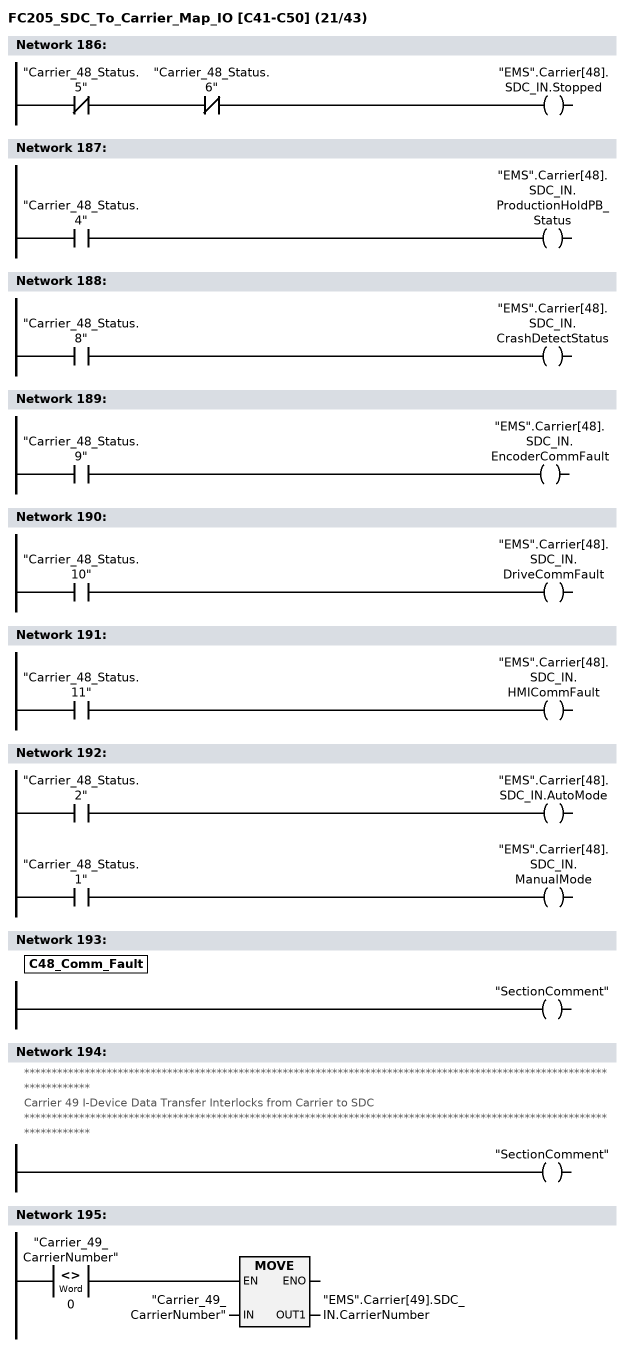
   RUNG wire#powerrail
      I_Contact( "Carrier_48_Status.5" )
      I_Contact( "Carrier_48_Status.6" )
      Coil( "EMS".Carrier[48].SDC_IN.Stopped )
   END_RUNG
   // the same network as SCL:
   "EMS".Carrier[48].SDC_IN.Stopped := NOT "Carrier_48_Status.5" AND NOT "Carrier_48_Status.6";
END_REGION

REGION Network 187
   RUNG wire#powerrail
      Contact( "Carrier_48_Status.4" )
      Coil( "EMS".Carrier[48].SDC_IN.ProductionHoldPB_Status )
   END_RUNG
   // the same network as SCL:
   "EMS".Carrier[48].SDC_IN.ProductionHoldPB_Status := "Carrier_48_Status.4";
END_REGION

REGION Network 188
   RUNG wire#powerrail
      Contact( "Carrier_48_Status.8" )
      Coil( "EMS".Carrier[48].SDC_IN.CrashDetectStatus )
   END_RUNG
   // the same network as SCL:
   "EMS".Carrier[48].SDC_IN.CrashDetectStatus := "Carrier_48_Status.8";
END_REGION

REGION Network 189
   RUNG wire#powerrail
      Contact( "Carrier_48_Status.9" )
      Coil( "EMS".Carrier[48].SDC_IN.EncoderCommFault )
   END_RUNG
   // the same network as SCL:
   "EMS".Carrier[48].SDC_IN.EncoderCommFault := "Carrier_48_Status.9";
END_REGION

REGION Network 190
   RUNG wire#powerrail
      Contact( "Carrier_48_Status.10" )
      Coil( "EMS".Carrier[48].SDC_IN.DriveCommFault )
   END_RUNG
   // the same network as SCL:
   "EMS".Carrier[48].SDC_IN.DriveCommFault := "Carrier_48_Status.10";
END_REGION

REGION Network 191
   RUNG wire#powerrail
      Contact( "Carrier_48_Status.11" )
      Coil( "EMS".Carrier[48].SDC_IN.HMICommFault )
   END_RUNG
   // the same network as SCL:
   "EMS".Carrier[48].SDC_IN.HMICommFault := "Carrier_48_Status.11";
END_REGION

REGION Network 192
   RUNG wire#powerrail
      Contact( "Carrier_48_Status.2" )
      Coil( "EMS".Carrier[48].SDC_IN.AutoMode )
   END_RUNG
   RUNG wire#powerrail
      Contact( "Carrier_48_Status.1" )
      Coil( "EMS".Carrier[48].SDC_IN.ManualMode )
   END_RUNG
   // the same network as SCL:
   "EMS".Carrier[48].SDC_IN.AutoMode := "Carrier_48_Status.2";
   "EMS".Carrier[48].SDC_IN.ManualMode := "Carrier_48_Status.1";
END_REGION

REGION Network 193
   Label( C48_Comm_Fault )
   RUNG wire#powerrail
      Coil( "SectionComment" )
   END_RUNG
   // the same network as SCL:
   C48_Comm_Fault:
   "SectionComment" := TRUE;
END_REGION

REGION Network 194
   // **********************************************************************************************************************
   // 
   // Carrier 49 I-Device Data Transfer Interlocks from Carrier to SDC
   // 
   // **********************************************************************************************************************
   RUNG wire#powerrail
      Coil( "SectionComment" )
   END_RUNG
   // the same network as SCL:
   "SectionComment" := TRUE;
END_REGION

REGION Network 195
   RUNG wire#powerrail
      { S7_Templates := "SrcType := Word" } NE_Contact(in1 := "Carrier_49_CarrierNumber", in2 := 0)
      Move(in := "Carrier_49_CarrierNumber", out1 => "EMS".Carrier[49].SDC_IN.CarrierNumber)
   END_RUNG
   // the same network as SCL:
   IF "Carrier_49_CarrierNumber" <> 0 THEN
       "EMS".Carrier[49].SDC_IN.CarrierNumber := "Carrier_49_CarrierNumber";
   END_IF;
END_REGION

REGION Network 196
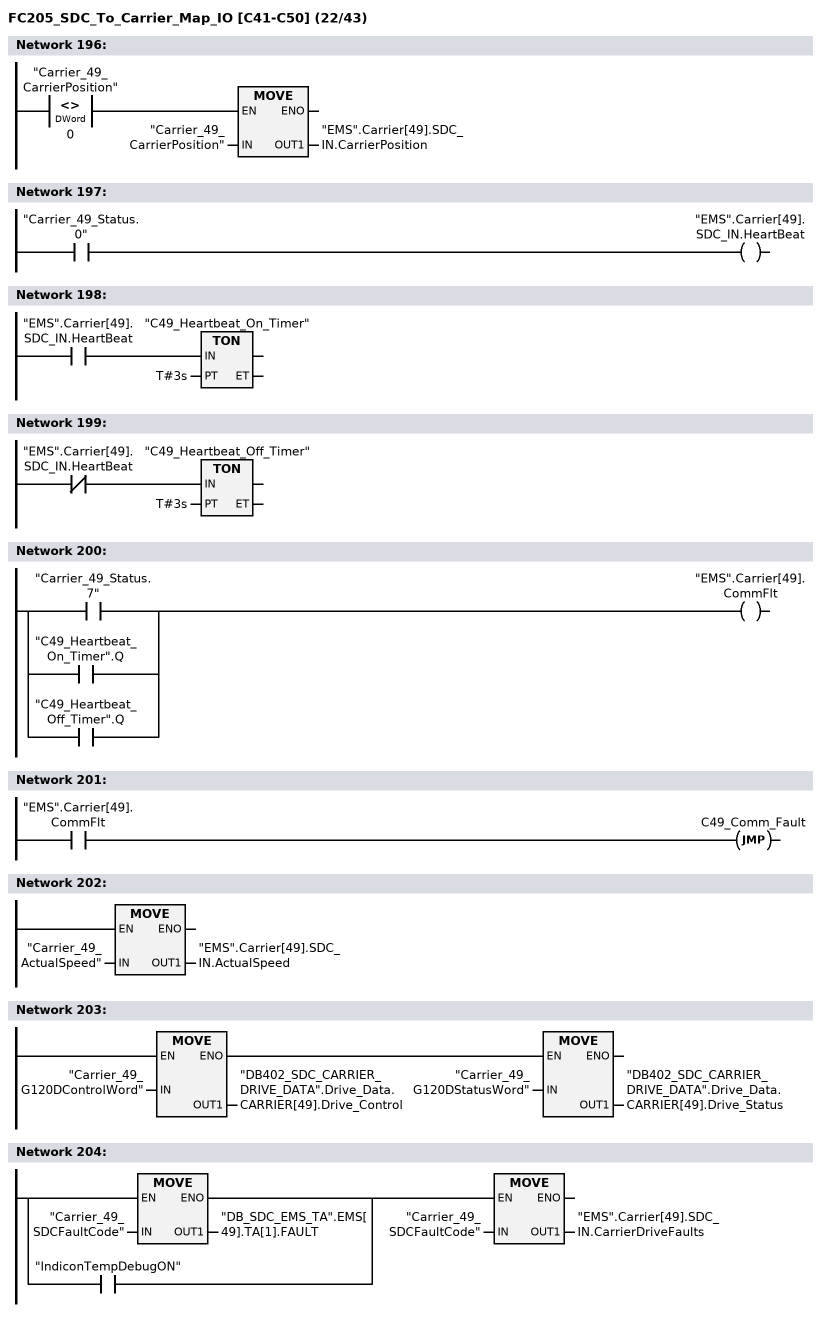
   RUNG wire#powerrail
      { S7_Templates := "SrcType := DWord" } NE_Contact(in1 := "Carrier_49_CarrierPosition", in2 := 0)
      Move(in := "Carrier_49_CarrierPosition", out1 => "EMS".Carrier[49].SDC_IN.CarrierPosition)
   END_RUNG
   // the same network as SCL:
   IF "Carrier_49_CarrierPosition" <> 0 THEN
       "EMS".Carrier[49].SDC_IN.CarrierPosition := "Carrier_49_CarrierPosition";
   END_IF;
END_REGION

REGION Network 197
   RUNG wire#powerrail
      Contact( "Carrier_49_Status.0" )
      Coil( "EMS".Carrier[49].SDC_IN.HeartBeat )
   END_RUNG
   // the same network as SCL:
   "EMS".Carrier[49].SDC_IN.HeartBeat := "Carrier_49_Status.0";
END_REGION

REGION Network 198
   "C49_Heartbeat_On_Timer".TON(IN := "EMS".Carrier[49].SDC_IN.HeartBeat, PT := T#3s);
END_REGION

REGION Network 199
   "C49_Heartbeat_Off_Timer".TON(IN := NOT "EMS".Carrier[49].SDC_IN.HeartBeat, PT := T#3s);
END_REGION

REGION Network 200
   RUNG wire#powerrail
      Contact( "Carrier_49_Status.7" )
      wire#w1
      Coil( "EMS".Carrier[49].CommFlt )
   END_RUNG
   RUNG wire#powerrail
      Contact( "C49_Heartbeat_On_Timer".Q )
   END_RUNG wire#w1
   RUNG wire#powerrail
      Contact( "C49_Heartbeat_Off_Timer".Q )
   END_RUNG wire#w1
   // the same network as SCL:
   "EMS".Carrier[49].CommFlt := "Carrier_49_Status.7" OR "C49_Heartbeat_On_Timer".Q OR "C49_Heartbeat_Off_Timer".Q;
END_REGION

REGION Network 201
   RUNG wire#powerrail
      Contact( "EMS".Carrier[49].CommFlt )
      JumpCoil( C49_Comm_Fault )
   END_RUNG
   // the same network as SCL:
   IF "EMS".Carrier[49].CommFlt THEN GOTO C49_Comm_Fault; END_IF;
END_REGION

REGION Network 202
   RUNG wire#powerrail
      Move(in := "Carrier_49_ActualSpeed", out1 => "EMS".Carrier[49].SDC_IN.ActualSpeed)
   END_RUNG
   // the same network as SCL:
   "EMS".Carrier[49].SDC_IN.ActualSpeed := "Carrier_49_ActualSpeed";
END_REGION

REGION Network 203
   RUNG wire#powerrail
      Move(in := "Carrier_49_G120DControlWord", out1 => "DB402_SDC_CARRIER_DRIVE_DATA".Drive_Data.CARRIER[49].Drive_Control)
      Move(in := "Carrier_49_G120DStatusWord", out1 => "DB402_SDC_CARRIER_DRIVE_DATA".Drive_Data.CARRIER[49].Drive_Status)
   END_RUNG
   // the same network as SCL:
   "DB402_SDC_CARRIER_DRIVE_DATA".Drive_Data.CARRIER[49].Drive_Control := "Carrier_49_G120DControlWord";
   "DB402_SDC_CARRIER_DRIVE_DATA".Drive_Data.CARRIER[49].Drive_Status := "Carrier_49_G120DStatusWord";
END_REGION

REGION Network 204
   RUNG wire#powerrail
      Move(in := "Carrier_49_SDCFaultCode", out1 => "DB_SDC_EMS_TA".EMS[49].TA[1].FAULT)
      wire#w1
      Move(in := "Carrier_49_SDCFaultCode", out1 => "EMS".Carrier[49].SDC_IN.CarrierDriveFaults)
   END_RUNG
   RUNG wire#powerrail
      Contact( "IndiconTempDebugON" )
   END_RUNG wire#w1
   // the same network as SCL:
   "DB_SDC_EMS_TA".EMS[49].TA[1].FAULT := "Carrier_49_SDCFaultCode";
   IF TRUE OR "IndiconTempDebugON" THEN
       "EMS".Carrier[49].SDC_IN.CarrierDriveFaults := "Carrier_49_SDCFaultCode";
   END_IF;
END_REGION

REGION Network 205
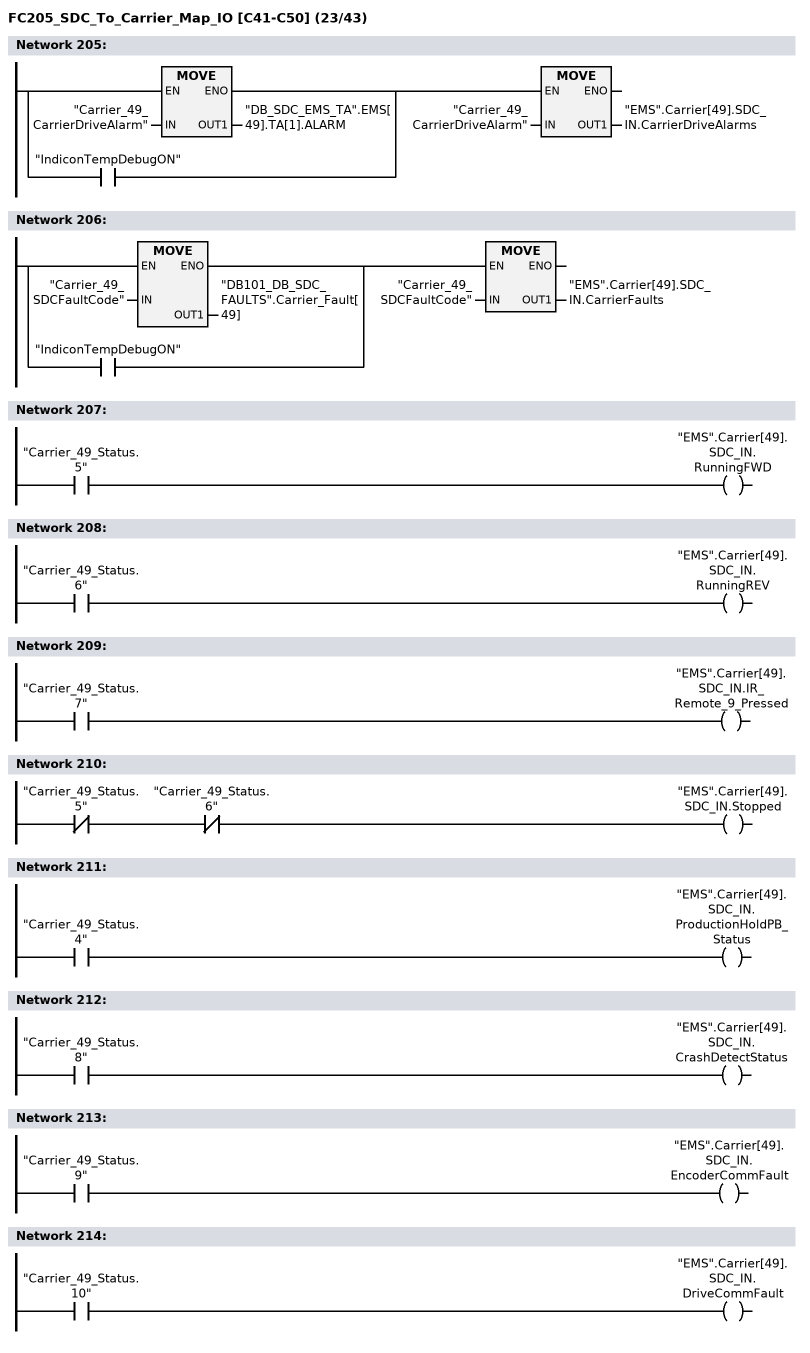
   RUNG wire#powerrail
      Move(in := "Carrier_49_CarrierDriveAlarm", out1 => "DB_SDC_EMS_TA".EMS[49].TA[1].ALARM)
      wire#w1
      Move(in := "Carrier_49_CarrierDriveAlarm", out1 => "EMS".Carrier[49].SDC_IN.CarrierDriveAlarms)
   END_RUNG
   RUNG wire#powerrail
      Contact( "IndiconTempDebugON" )
   END_RUNG wire#w1
   // the same network as SCL:
   "DB_SDC_EMS_TA".EMS[49].TA[1].ALARM := "Carrier_49_CarrierDriveAlarm";
   IF TRUE OR "IndiconTempDebugON" THEN
       "EMS".Carrier[49].SDC_IN.CarrierDriveAlarms := "Carrier_49_CarrierDriveAlarm";
   END_IF;
END_REGION

REGION Network 206
   RUNG wire#powerrail
      Move(in := "Carrier_49_SDCFaultCode", out1 => "DB101_DB_SDC_FAULTS".Carrier_Fault[49])
      wire#w1
      Move(in := "Carrier_49_SDCFaultCode", out1 => "EMS".Carrier[49].SDC_IN.CarrierFaults)
   END_RUNG
   RUNG wire#powerrail
      Contact( "IndiconTempDebugON" )
   END_RUNG wire#w1
   // the same network as SCL:
   "DB101_DB_SDC_FAULTS".Carrier_Fault[49] := "Carrier_49_SDCFaultCode";
   IF TRUE OR "IndiconTempDebugON" THEN
       "EMS".Carrier[49].SDC_IN.CarrierFaults := "Carrier_49_SDCFaultCode";
   END_IF;
END_REGION

REGION Network 207
   RUNG wire#powerrail
      Contact( "Carrier_49_Status.5" )
      Coil( "EMS".Carrier[49].SDC_IN.RunningFWD )
   END_RUNG
   // the same network as SCL:
   "EMS".Carrier[49].SDC_IN.RunningFWD := "Carrier_49_Status.5";
END_REGION

REGION Network 208
   RUNG wire#powerrail
      Contact( "Carrier_49_Status.6" )
      Coil( "EMS".Carrier[49].SDC_IN.RunningREV )
   END_RUNG
   // the same network as SCL:
   "EMS".Carrier[49].SDC_IN.RunningREV := "Carrier_49_Status.6";
END_REGION

REGION Network 209
   RUNG wire#powerrail
      Contact( "Carrier_49_Status.7" )
      Coil( "EMS".Carrier[49].SDC_IN.IR_Remote_9_Pressed )
   END_RUNG
   // the same network as SCL:
   "EMS".Carrier[49].SDC_IN.IR_Remote_9_Pressed := "Carrier_49_Status.7";
END_REGION

REGION Network 210
   RUNG wire#powerrail
      I_Contact( "Carrier_49_Status.5" )
      I_Contact( "Carrier_49_Status.6" )
      Coil( "EMS".Carrier[49].SDC_IN.Stopped )
   END_RUNG
   // the same network as SCL:
   "EMS".Carrier[49].SDC_IN.Stopped := NOT "Carrier_49_Status.5" AND NOT "Carrier_49_Status.6";
END_REGION

REGION Network 211
   RUNG wire#powerrail
      Contact( "Carrier_49_Status.4" )
      Coil( "EMS".Carrier[49].SDC_IN.ProductionHoldPB_Status )
   END_RUNG
   // the same network as SCL:
   "EMS".Carrier[49].SDC_IN.ProductionHoldPB_Status := "Carrier_49_Status.4";
END_REGION

REGION Network 212
   RUNG wire#powerrail
      Contact( "Carrier_49_Status.8" )
      Coil( "EMS".Carrier[49].SDC_IN.CrashDetectStatus )
   END_RUNG
   // the same network as SCL:
   "EMS".Carrier[49].SDC_IN.CrashDetectStatus := "Carrier_49_Status.8";
END_REGION

REGION Network 213
   RUNG wire#powerrail
      Contact( "Carrier_49_Status.9" )
      Coil( "EMS".Carrier[49].SDC_IN.EncoderCommFault )
   END_RUNG
   // the same network as SCL:
   "EMS".Carrier[49].SDC_IN.EncoderCommFault := "Carrier_49_Status.9";
END_REGION

REGION Network 214
   RUNG wire#powerrail
      Contact( "Carrier_49_Status.10" )
      Coil( "EMS".Carrier[49].SDC_IN.DriveCommFault )
   END_RUNG
   // the same network as SCL:
   "EMS".Carrier[49].SDC_IN.DriveCommFault := "Carrier_49_Status.10";
END_REGION

REGION Network 215
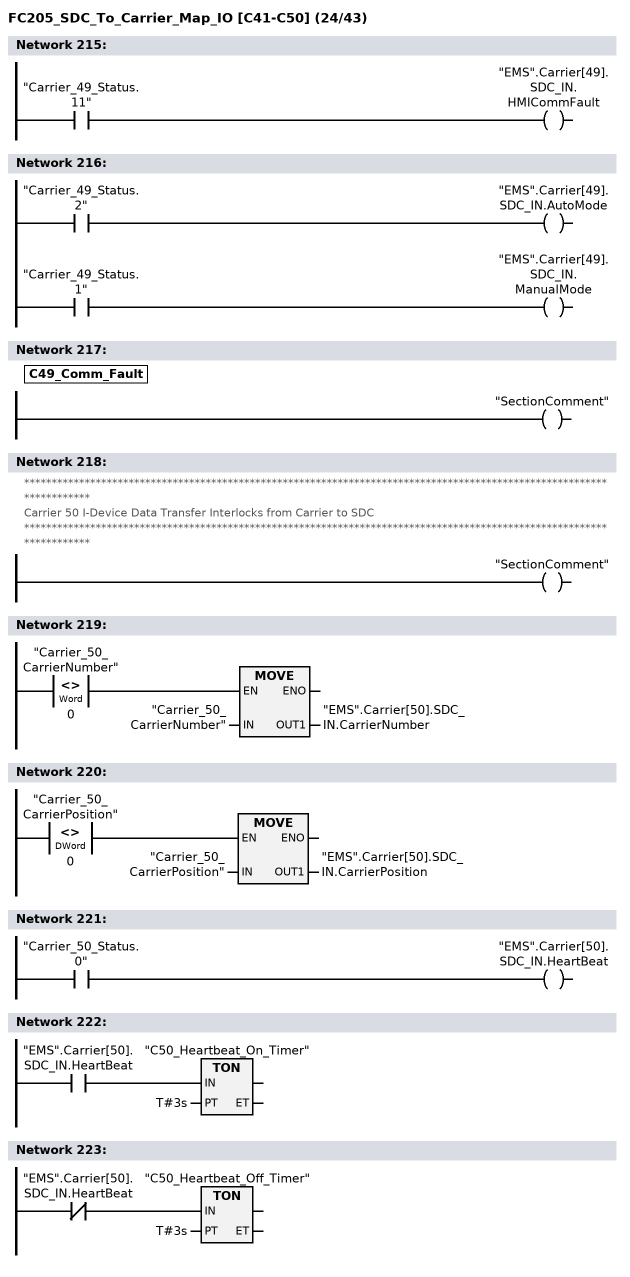
   RUNG wire#powerrail
      Contact( "Carrier_49_Status.11" )
      Coil( "EMS".Carrier[49].SDC_IN.HMICommFault )
   END_RUNG
   // the same network as SCL:
   "EMS".Carrier[49].SDC_IN.HMICommFault := "Carrier_49_Status.11";
END_REGION

REGION Network 216
   RUNG wire#powerrail
      Contact( "Carrier_49_Status.2" )
      Coil( "EMS".Carrier[49].SDC_IN.AutoMode )
   END_RUNG
   RUNG wire#powerrail
      Contact( "Carrier_49_Status.1" )
      Coil( "EMS".Carrier[49].SDC_IN.ManualMode )
   END_RUNG
   // the same network as SCL:
   "EMS".Carrier[49].SDC_IN.AutoMode := "Carrier_49_Status.2";
   "EMS".Carrier[49].SDC_IN.ManualMode := "Carrier_49_Status.1";
END_REGION

REGION Network 217
   Label( C49_Comm_Fault )
   RUNG wire#powerrail
      Coil( "SectionComment" )
   END_RUNG
   // the same network as SCL:
   C49_Comm_Fault:
   "SectionComment" := TRUE;
END_REGION

REGION Network 218
   // **********************************************************************************************************************
   // 
   // Carrier 50 I-Device Data Transfer Interlocks from Carrier to SDC
   // 
   // **********************************************************************************************************************
   RUNG wire#powerrail
      Coil( "SectionComment" )
   END_RUNG
   // the same network as SCL:
   "SectionComment" := TRUE;
END_REGION

REGION Network 219
   RUNG wire#powerrail
      { S7_Templates := "SrcType := Word" } NE_Contact(in1 := "Carrier_50_CarrierNumber", in2 := 0)
      Move(in := "Carrier_50_CarrierNumber", out1 => "EMS".Carrier[50].SDC_IN.CarrierNumber)
   END_RUNG
   // the same network as SCL:
   IF "Carrier_50_CarrierNumber" <> 0 THEN
       "EMS".Carrier[50].SDC_IN.CarrierNumber := "Carrier_50_CarrierNumber";
   END_IF;
END_REGION

REGION Network 220
   RUNG wire#powerrail
      { S7_Templates := "SrcType := DWord" } NE_Contact(in1 := "Carrier_50_CarrierPosition", in2 := 0)
      Move(in := "Carrier_50_CarrierPosition", out1 => "EMS".Carrier[50].SDC_IN.CarrierPosition)
   END_RUNG
   // the same network as SCL:
   IF "Carrier_50_CarrierPosition" <> 0 THEN
       "EMS".Carrier[50].SDC_IN.CarrierPosition := "Carrier_50_CarrierPosition";
   END_IF;
END_REGION

REGION Network 221
   RUNG wire#powerrail
      Contact( "Carrier_50_Status.0" )
      Coil( "EMS".Carrier[50].SDC_IN.HeartBeat )
   END_RUNG
   // the same network as SCL:
   "EMS".Carrier[50].SDC_IN.HeartBeat := "Carrier_50_Status.0";
END_REGION

REGION Network 222
   "C50_Heartbeat_On_Timer".TON(IN := "EMS".Carrier[50].SDC_IN.HeartBeat, PT := T#3s);
END_REGION

REGION Network 223
   "C50_Heartbeat_Off_Timer".TON(IN := NOT "EMS".Carrier[50].SDC_IN.HeartBeat, PT := T#3s);
END_REGION

REGION Network 224
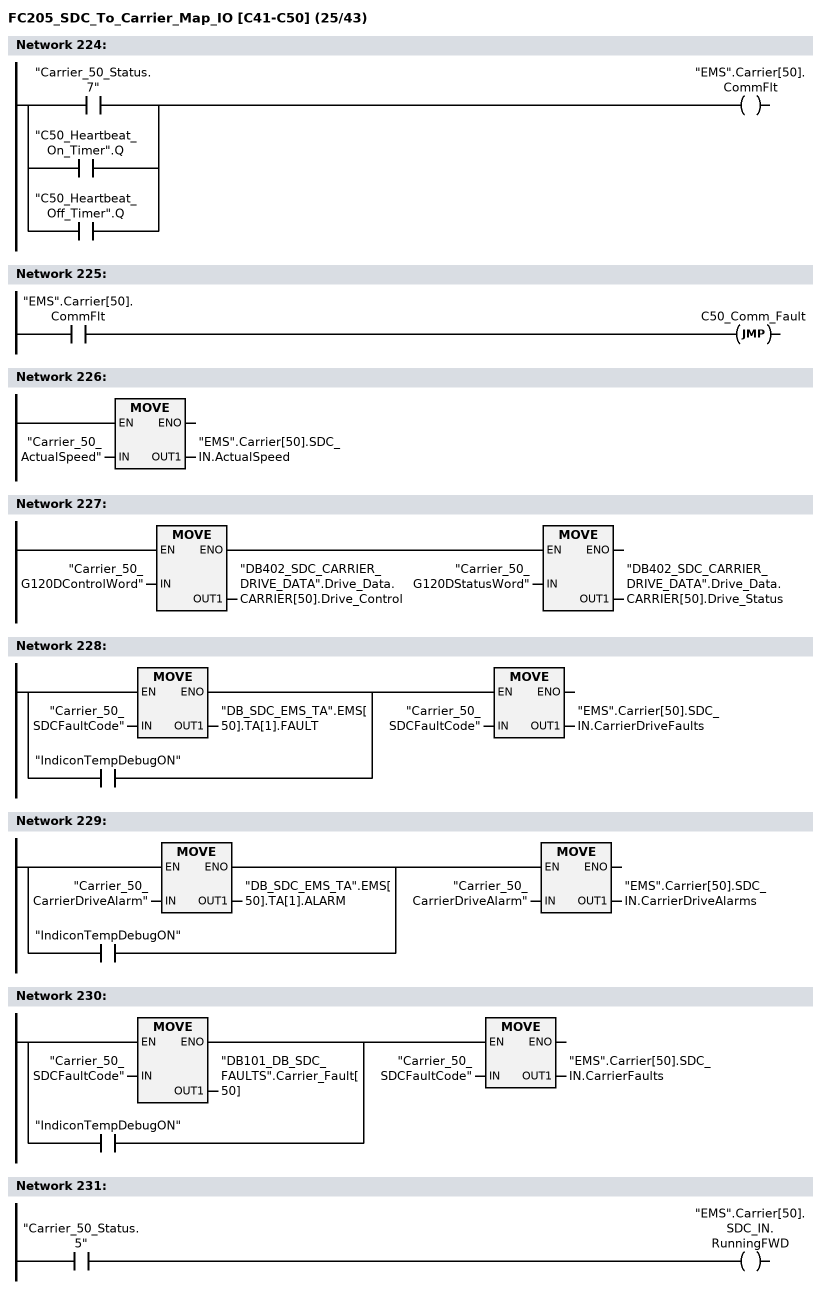
   RUNG wire#powerrail
      Contact( "Carrier_50_Status.7" )
      wire#w1
      Coil( "EMS".Carrier[50].CommFlt )
   END_RUNG
   RUNG wire#powerrail
      Contact( "C50_Heartbeat_On_Timer".Q )
   END_RUNG wire#w1
   RUNG wire#powerrail
      Contact( "C50_Heartbeat_Off_Timer".Q )
   END_RUNG wire#w1
   // the same network as SCL:
   "EMS".Carrier[50].CommFlt := "Carrier_50_Status.7" OR "C50_Heartbeat_On_Timer".Q OR "C50_Heartbeat_Off_Timer".Q;
END_REGION

REGION Network 225
   RUNG wire#powerrail
      Contact( "EMS".Carrier[50].CommFlt )
      JumpCoil( C50_Comm_Fault )
   END_RUNG
   // the same network as SCL:
   IF "EMS".Carrier[50].CommFlt THEN GOTO C50_Comm_Fault; END_IF;
END_REGION

REGION Network 226
   RUNG wire#powerrail
      Move(in := "Carrier_50_ActualSpeed", out1 => "EMS".Carrier[50].SDC_IN.ActualSpeed)
   END_RUNG
   // the same network as SCL:
   "EMS".Carrier[50].SDC_IN.ActualSpeed := "Carrier_50_ActualSpeed";
END_REGION

REGION Network 227
   RUNG wire#powerrail
      Move(in := "Carrier_50_G120DControlWord", out1 => "DB402_SDC_CARRIER_DRIVE_DATA".Drive_Data.CARRIER[50].Drive_Control)
      Move(in := "Carrier_50_G120DStatusWord", out1 => "DB402_SDC_CARRIER_DRIVE_DATA".Drive_Data.CARRIER[50].Drive_Status)
   END_RUNG
   // the same network as SCL:
   "DB402_SDC_CARRIER_DRIVE_DATA".Drive_Data.CARRIER[50].Drive_Control := "Carrier_50_G120DControlWord";
   "DB402_SDC_CARRIER_DRIVE_DATA".Drive_Data.CARRIER[50].Drive_Status := "Carrier_50_G120DStatusWord";
END_REGION

REGION Network 228
   RUNG wire#powerrail
      Move(in := "Carrier_50_SDCFaultCode", out1 => "DB_SDC_EMS_TA".EMS[50].TA[1].FAULT)
      wire#w1
      Move(in := "Carrier_50_SDCFaultCode", out1 => "EMS".Carrier[50].SDC_IN.CarrierDriveFaults)
   END_RUNG
   RUNG wire#powerrail
      Contact( "IndiconTempDebugON" )
   END_RUNG wire#w1
   // the same network as SCL:
   "DB_SDC_EMS_TA".EMS[50].TA[1].FAULT := "Carrier_50_SDCFaultCode";
   IF TRUE OR "IndiconTempDebugON" THEN
       "EMS".Carrier[50].SDC_IN.CarrierDriveFaults := "Carrier_50_SDCFaultCode";
   END_IF;
END_REGION

REGION Network 229
   RUNG wire#powerrail
      Move(in := "Carrier_50_CarrierDriveAlarm", out1 => "DB_SDC_EMS_TA".EMS[50].TA[1].ALARM)
      wire#w1
      Move(in := "Carrier_50_CarrierDriveAlarm", out1 => "EMS".Carrier[50].SDC_IN.CarrierDriveAlarms)
   END_RUNG
   RUNG wire#powerrail
      Contact( "IndiconTempDebugON" )
   END_RUNG wire#w1
   // the same network as SCL:
   "DB_SDC_EMS_TA".EMS[50].TA[1].ALARM := "Carrier_50_CarrierDriveAlarm";
   IF TRUE OR "IndiconTempDebugON" THEN
       "EMS".Carrier[50].SDC_IN.CarrierDriveAlarms := "Carrier_50_CarrierDriveAlarm";
   END_IF;
END_REGION

REGION Network 230
   RUNG wire#powerrail
      Move(in := "Carrier_50_SDCFaultCode", out1 => "DB101_DB_SDC_FAULTS".Carrier_Fault[50])
      wire#w1
      Move(in := "Carrier_50_SDCFaultCode", out1 => "EMS".Carrier[50].SDC_IN.CarrierFaults)
   END_RUNG
   RUNG wire#powerrail
      Contact( "IndiconTempDebugON" )
   END_RUNG wire#w1
   // the same network as SCL:
   "DB101_DB_SDC_FAULTS".Carrier_Fault[50] := "Carrier_50_SDCFaultCode";
   IF TRUE OR "IndiconTempDebugON" THEN
       "EMS".Carrier[50].SDC_IN.CarrierFaults := "Carrier_50_SDCFaultCode";
   END_IF;
END_REGION

REGION Network 231
   RUNG wire#powerrail
      Contact( "Carrier_50_Status.5" )
      Coil( "EMS".Carrier[50].SDC_IN.RunningFWD )
   END_RUNG
   // the same network as SCL:
   "EMS".Carrier[50].SDC_IN.RunningFWD := "Carrier_50_Status.5";
END_REGION

REGION Network 232
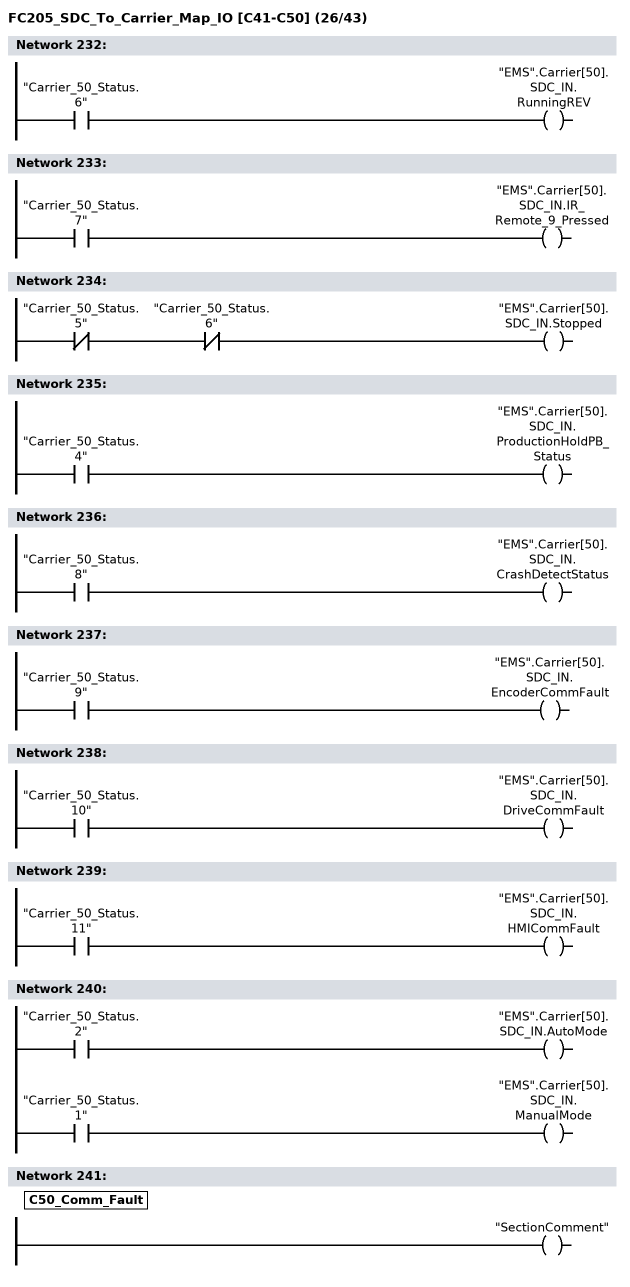
   RUNG wire#powerrail
      Contact( "Carrier_50_Status.6" )
      Coil( "EMS".Carrier[50].SDC_IN.RunningREV )
   END_RUNG
   // the same network as SCL:
   "EMS".Carrier[50].SDC_IN.RunningREV := "Carrier_50_Status.6";
END_REGION

REGION Network 233
   RUNG wire#powerrail
      Contact( "Carrier_50_Status.7" )
      Coil( "EMS".Carrier[50].SDC_IN.IR_Remote_9_Pressed )
   END_RUNG
   // the same network as SCL:
   "EMS".Carrier[50].SDC_IN.IR_Remote_9_Pressed := "Carrier_50_Status.7";
END_REGION

REGION Network 234
   RUNG wire#powerrail
      I_Contact( "Carrier_50_Status.5" )
      I_Contact( "Carrier_50_Status.6" )
      Coil( "EMS".Carrier[50].SDC_IN.Stopped )
   END_RUNG
   // the same network as SCL:
   "EMS".Carrier[50].SDC_IN.Stopped := NOT "Carrier_50_Status.5" AND NOT "Carrier_50_Status.6";
END_REGION

REGION Network 235
   RUNG wire#powerrail
      Contact( "Carrier_50_Status.4" )
      Coil( "EMS".Carrier[50].SDC_IN.ProductionHoldPB_Status )
   END_RUNG
   // the same network as SCL:
   "EMS".Carrier[50].SDC_IN.ProductionHoldPB_Status := "Carrier_50_Status.4";
END_REGION

REGION Network 236
   RUNG wire#powerrail
      Contact( "Carrier_50_Status.8" )
      Coil( "EMS".Carrier[50].SDC_IN.CrashDetectStatus )
   END_RUNG
   // the same network as SCL:
   "EMS".Carrier[50].SDC_IN.CrashDetectStatus := "Carrier_50_Status.8";
END_REGION

REGION Network 237
   RUNG wire#powerrail
      Contact( "Carrier_50_Status.9" )
      Coil( "EMS".Carrier[50].SDC_IN.EncoderCommFault )
   END_RUNG
   // the same network as SCL:
   "EMS".Carrier[50].SDC_IN.EncoderCommFault := "Carrier_50_Status.9";
END_REGION

REGION Network 238
   RUNG wire#powerrail
      Contact( "Carrier_50_Status.10" )
      Coil( "EMS".Carrier[50].SDC_IN.DriveCommFault )
   END_RUNG
   // the same network as SCL:
   "EMS".Carrier[50].SDC_IN.DriveCommFault := "Carrier_50_Status.10";
END_REGION

REGION Network 239
   RUNG wire#powerrail
      Contact( "Carrier_50_Status.11" )
      Coil( "EMS".Carrier[50].SDC_IN.HMICommFault )
   END_RUNG
   // the same network as SCL:
   "EMS".Carrier[50].SDC_IN.HMICommFault := "Carrier_50_Status.11";
END_REGION

REGION Network 240
   RUNG wire#powerrail
      Contact( "Carrier_50_Status.2" )
      Coil( "EMS".Carrier[50].SDC_IN.AutoMode )
   END_RUNG
   RUNG wire#powerrail
      Contact( "Carrier_50_Status.1" )
      Coil( "EMS".Carrier[50].SDC_IN.ManualMode )
   END_RUNG
   // the same network as SCL:
   "EMS".Carrier[50].SDC_IN.AutoMode := "Carrier_50_Status.2";
   "EMS".Carrier[50].SDC_IN.ManualMode := "Carrier_50_Status.1";
END_REGION

REGION Network 241
   Label( C50_Comm_Fault )
   RUNG wire#powerrail
      Coil( "SectionComment" )
   END_RUNG
   // the same network as SCL:
   C50_Comm_Fault:
   "SectionComment" := TRUE;
END_REGION

REGION Network 242
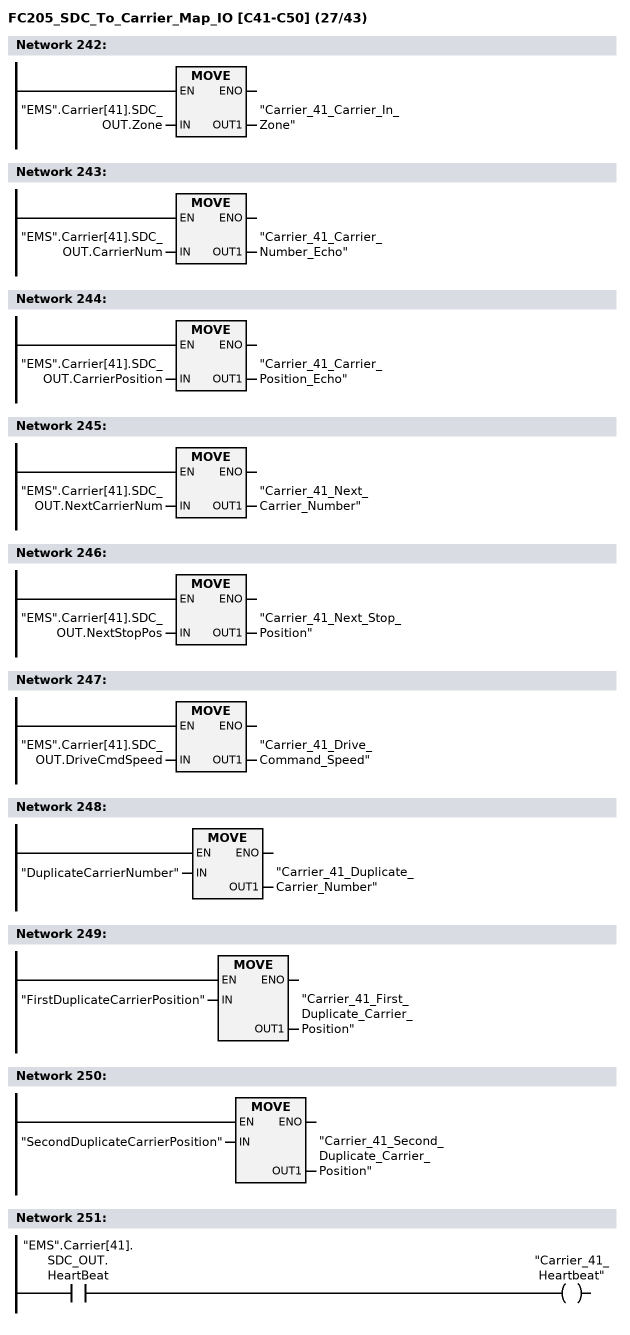
   RUNG wire#powerrail
      Move(in := "EMS".Carrier[41].SDC_OUT.Zone, out1 => "Carrier_41_Carrier_In_Zone")
   END_RUNG
   // the same network as SCL:
   "Carrier_41_Carrier_In_Zone" := "EMS".Carrier[41].SDC_OUT.Zone;
END_REGION

REGION Network 243
   RUNG wire#powerrail
      Move(in := "EMS".Carrier[41].SDC_OUT.CarrierNum, out1 => "Carrier_41_Carrier_Number_Echo")
   END_RUNG
   // the same network as SCL:
   "Carrier_41_Carrier_Number_Echo" := "EMS".Carrier[41].SDC_OUT.CarrierNum;
END_REGION

REGION Network 244
   RUNG wire#powerrail
      Move(in := "EMS".Carrier[41].SDC_OUT.CarrierPosition, out1 => "Carrier_41_Carrier_Position_Echo")
   END_RUNG
   // the same network as SCL:
   "Carrier_41_Carrier_Position_Echo" := "EMS".Carrier[41].SDC_OUT.CarrierPosition;
END_REGION

REGION Network 245
   RUNG wire#powerrail
      Move(in := "EMS".Carrier[41].SDC_OUT.NextCarrierNum, out1 => "Carrier_41_Next_Carrier_Number")
   END_RUNG
   // the same network as SCL:
   "Carrier_41_Next_Carrier_Number" := "EMS".Carrier[41].SDC_OUT.NextCarrierNum;
END_REGION

REGION Network 246
   RUNG wire#powerrail
      Move(in := "EMS".Carrier[41].SDC_OUT.NextStopPos, out1 => "Carrier_41_Next_Stop_Position")
   END_RUNG
   // the same network as SCL:
   "Carrier_41_Next_Stop_Position" := "EMS".Carrier[41].SDC_OUT.NextStopPos;
END_REGION

REGION Network 247
   RUNG wire#powerrail
      Move(in := "EMS".Carrier[41].SDC_OUT.DriveCmdSpeed, out1 => "Carrier_41_Drive_Command_Speed")
   END_RUNG
   // the same network as SCL:
   "Carrier_41_Drive_Command_Speed" := "EMS".Carrier[41].SDC_OUT.DriveCmdSpeed;
END_REGION

REGION Network 248
   RUNG wire#powerrail
      Move(in := "DuplicateCarrierNumber", out1 => "Carrier_41_Duplicate_Carrier_Number")
   END_RUNG
   // the same network as SCL:
   "Carrier_41_Duplicate_Carrier_Number" := "DuplicateCarrierNumber";
END_REGION

REGION Network 249
   RUNG wire#powerrail
      Move(in := "FirstDuplicateCarrierPosition", out1 => "Carrier_41_First_Duplicate_Carrier_Position")
   END_RUNG
   // the same network as SCL:
   "Carrier_41_First_Duplicate_Carrier_Position" := "FirstDuplicateCarrierPosition";
END_REGION

REGION Network 250
   RUNG wire#powerrail
      Move(in := "SecondDuplicateCarrierPosition", out1 => "Carrier_41_Second_Duplicate_Carrier_Position")
   END_RUNG
   // the same network as SCL:
   "Carrier_41_Second_Duplicate_Carrier_Position" := "SecondDuplicateCarrierPosition";
END_REGION

REGION Network 251
   RUNG wire#powerrail
      Contact( "EMS".Carrier[41].SDC_OUT.HeartBeat )
      Coil( "Carrier_41_Heartbeat" )
   END_RUNG
   // the same network as SCL:
   "Carrier_41_Heartbeat" := "EMS".Carrier[41].SDC_OUT.HeartBeat;
END_REGION

REGION Network 252
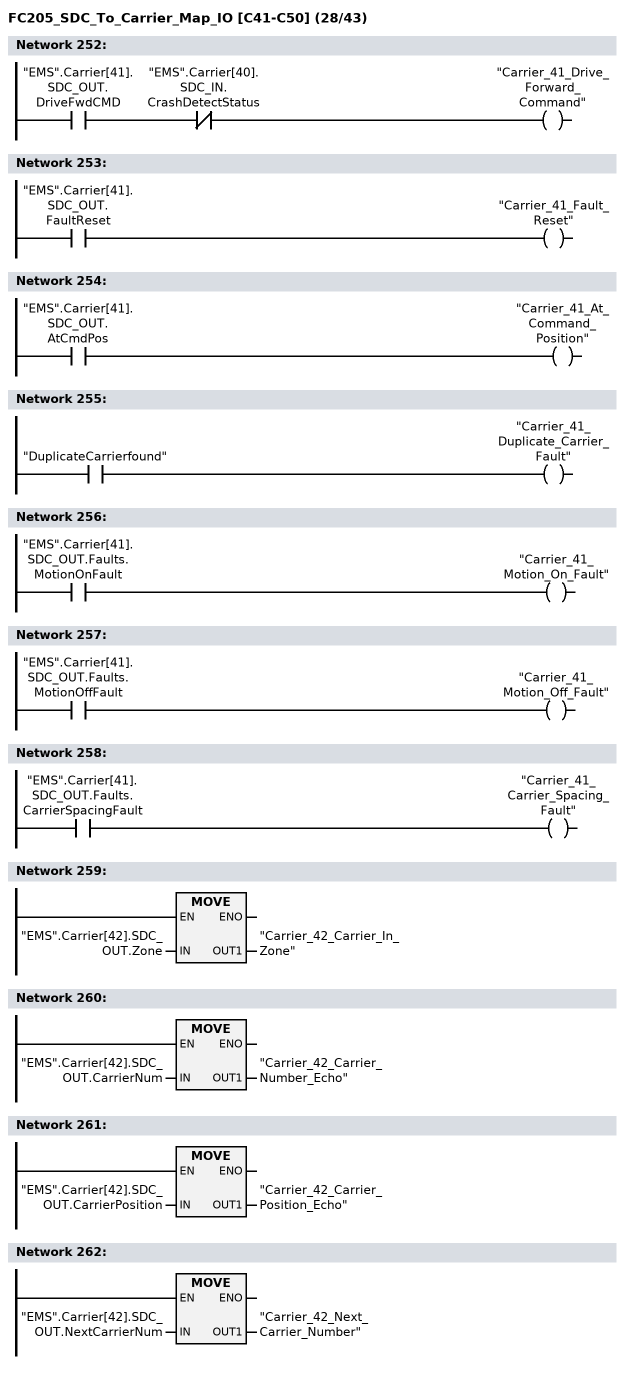
   RUNG wire#powerrail
      Contact( "EMS".Carrier[41].SDC_OUT.DriveFwdCMD )
      I_Contact( "EMS".Carrier[40].SDC_IN.CrashDetectStatus )
      Coil( "Carrier_41_Drive_Forward_Command" )
   END_RUNG
   // the same network as SCL:
   "Carrier_41_Drive_Forward_Command" := "EMS".Carrier[41].SDC_OUT.DriveFwdCMD AND NOT "EMS".Carrier[40].SDC_IN.CrashDetectStatus;
END_REGION

REGION Network 253
   RUNG wire#powerrail
      Contact( "EMS".Carrier[41].SDC_OUT.FaultReset )
      Coil( "Carrier_41_Fault_Reset" )
   END_RUNG
   // the same network as SCL:
   "Carrier_41_Fault_Reset" := "EMS".Carrier[41].SDC_OUT.FaultReset;
END_REGION

REGION Network 254
   RUNG wire#powerrail
      Contact( "EMS".Carrier[41].SDC_OUT.AtCmdPos )
      Coil( "Carrier_41_At_Command_Position" )
   END_RUNG
   // the same network as SCL:
   "Carrier_41_At_Command_Position" := "EMS".Carrier[41].SDC_OUT.AtCmdPos;
END_REGION

REGION Network 255
   RUNG wire#powerrail
      Contact( "DuplicateCarrierfound" )
      Coil( "Carrier_41_Duplicate_Carrier_Fault" )
   END_RUNG
   // the same network as SCL:
   "Carrier_41_Duplicate_Carrier_Fault" := "DuplicateCarrierfound";
END_REGION
